screen "eProC - 09 - Estados PL_Diag" 1280x770, template "Template"
   Rectangle "Rectángulo_1" at 146,344 size 393x149
      Visibility <- "STOP_RUN"
   Button "Botón_2" at 352,429 size 144x40; TextOff 'Reset'
      on Click: SetBit("PL_Reset")
      Visibility <- "STOP_RUN"
   Button "Botón_1" at 192,429 size 144x40; TextOff 'Continuar'
      on Click: SetBit("PL_Continuar")
      Visibility <- "STOP_RUN"
   TextField "Campo de texto_17" at 165,356 size 351x73; Text 'Se ha detectado un reinicio del PLC. ¿Qué desea hacer con el ciclo de la Plegadora?'
      Visibility <- "STOP_RUN"
   Rectangle "Rectángulo_13" at 687,65 size 29x579
      Visibility <- "PL_S_1"
   Rectangle "Rectángulo_15" at 727,65 size 29x579
      Visibility <- "PL_S_2"
   Rectangle "Rectángulo_16" at 767,65 size 29x579
      Visibility <- "PL_S_9"
   Rectangle "Rectángulo_17" at 807,65 size 29x579
      Visibility <- "PL_S_3"
   Rectangle "Rectángulo_18" at 847,65 size 29x579
      Visibility <- "PL_S_4"
   Rectangle "Rectángulo_19" at 887,65 size 29x579
      Visibility <- "PL_S_10"
   Rectangle "Rectángulo_20" at 927,65 size 29x579
      Visibility <- "PL_S_5"
   Rectangle "Rectángulo_21" at 967,65 size 29x579
      Visibility <- "PL_S_11"
   Rectangle "Rectángulo_22" at 1007,65 size 29x579
      Visibility <- "PL_S_6"
   Rectangle "Rectángulo_23" at 647,65 size 29x579
      Visibility <- "PL_S_12"
   Circle "Círculo_2" at 78,143 size 450x450
      Appearance <- "PL_en_Ciclo"
   SymbolicIOField "Campo ES simbólico_1" at 109,310 size 387x69; TextOn '1'; TextOff '0'; TextList "Estados_PL"
      ProcessValue <- "PL_Estados"
   Polygon "Polígono_1" at 466,215 size 12x13
      Appearance <- "PL_en_Ciclo"
   Polygon "Polígono_2" at 520,333 size 8x12
      Appearance <- "PL_en_Ciclo"
   Polygon "Polígono_3" at 503,456 size 8x12
      Appearance <- "PL_en_Ciclo"
   Polygon "Polígono_4" at 401,559 size 14x10
      Appearance <- "PL_en_Ciclo"
   Polygon "Polígono_5" at 242,583 size 14x7
      Appearance <- "PL_en_Ciclo"
   Polygon "Polígono_6" at 124,503 size 10x13
      Appearance <- "PL_en_Ciclo"
   Polygon "Polígono_7" at 78,389 size 6x17
      Appearance <- "PL_en_Ciclo"
   Polygon "Polígono_8" at 94,269 size 7x14
      Appearance <- "PL_en_Ciclo"
   Polygon "Polígono_9" at 345,145 size 13x6
      Appearance <- "PL_en_Ciclo"
   Polygon "Polígono_10" at 186,169 size 12x9
      Appearance <- "PL_en_Ciclo"
   GraphicIOField "Campo ES gráfico_1" at 90,461 size 50x46; PictureList "Estado"
      ProcessValue <- "PL_S_11"
   GraphicIOField "Campo ES gráfico_2" at 55,345 size 50x46; PictureList "Estado"
      ProcessValue <- "PL_S_6"
   GraphicIOField "Campo ES gráfico_4" at 196,137 size 50x46; PictureList "Estado"
      ProcessValue <- "PL_S_1"
   GraphicIOField "Campo ES gráfico_5" at 196,555 size 50x46; PictureList "Estado"
      ProcessValue <- "PL_S_5"
   GraphicIOField "Campo ES gráfico_6" at 356,137 size 50x46; PictureList "Estado"
      ProcessValue <- "PL_S_2"
   GraphicIOField "Campo ES gráfico_7" at 356,554 size 50x46; PictureList "Estado"
      ProcessValue <- "PL_S_10"
   GraphicIOField "Campo ES gráfico_8" at 467,464 size 50x46; PictureList "Estado"
      ProcessValue <- "PL_S_4"
   GraphicIOField "Campo ES gráfico_9" at 466,226 size 50x46; PictureList "Estado"
      ProcessValue <- "PL_S_9"
   GraphicIOField "Campo ES gráfico_10" at 501,345 size 50x46; PictureList "Estado"
      ProcessValue <- "PL_S_3"
   SymbolicIOField "Campo ES simbólico_2" at 103,359 size 403x45; TextOn '1'; TextOff '0'; TextList "Transiciones_PL"
      ProcessValue <- "PL_Estados"
   Line "Línea_1" at 109,126 size 0x102
      Appearance <- "PL_en_Ciclo"
   Polygon "Polígono_11" at 106,213 size 7x15
      Appearance <- "PL_en_Ciclo"
   GraphicIOField "Campo ES gráfico_11" at 84,121 size 50x46; PictureList "Estado"
      ProcessValue <- "PL_S_0"
   GraphicIOField "Campo ES gráfico_3" at 86,226 size 50x46; PictureList "Estado"
      ProcessValue <- "PL_S_12"
   TextField "Campo de texto_1" at 31,36 size 300x29; Text 'Máquina de estados Plegadores'
   TextField "Campo de texto_15" at 372,147 size 16x25; Text '2'
   TextField "Campo de texto_16" at 482,236 size 16x25; Text '9'
   TextField "Campo de texto_13" at 518,355 size 16x25; Text '3'
   TextField "Campo de texto_24" at 483,474 size 16x25; Text '4'
   TextField "Campo de texto_26" at 366,564 size 30x25; Text '10'
   TextField "Campo de texto_27" at 211,565 size 19x25; Text '5'
   TextField "Campo de texto_28" at 100,471 size 30x25; Text '11'
   TextField "Campo de texto_29" at 70,355 size 15x25; Text '6'
   TextField "Campo de texto_30" at 96,236 size 31x25; Text '12'
   TextField "Campo de texto_31" at 212,147 size 16x25; Text '1'
   TextField "Campo de texto_32" at 100,131 size 16x25; Text '0'
   TextField "Campo de texto_2" at 1101,68 size 42x21; Text 'M10.3'
   TextField "Campo de texto_3" at 1147,92 size 50x21; Text 'M180.0'
   TextField "Campo de texto_4" at 1145,116 size 50x21; Text 'M180.1'
   TextField "Campo de texto_5" at 1170,140 size 50x21; Text 'M180.3'
   TextField "Campo de texto_6" at 1176,164 size 50x21; Text 'M180.4'
   TextField "Campo de texto_8" at 1138,212 size 96x21; Text 'DB11.DBX46.0'
   TextField "Campo de texto_14" at 1134,500 size 50x21; Text 'M170.5'
   TextField "Campo de texto_7" at 1134,524 size 50x21; Text 'M170.6'
   TextField "Campo de texto_9" at 1140,548 size 50x21; Text 'M170.7'
   TextField "Campo de texto_10" at 1147,572 size 50x21; Text 'M171.0'
   TextField "Campo de texto_11" at 1149,596 size 50x21; Text 'M171.1'
   TextField "Campo de texto_18" at 1130,620 size 50x21; Text 'M171.2'
   TextField "Campo de texto_22" at 1141,260 size 50x21; Text 'M165.0'
   TextField "Campo de texto_23" at 1148,284 size 50x21; Text 'M165.1'
   TextField "Campo de texto_12" at 1119,308 size 50x21; Text 'M165.2'
   TextField "Campo de texto_25" at 1125,332 size 50x21; Text 'M165.3'
   TextField "Campo de texto_19" at 1121,356 size 50x21; Text 'M165.4'
   TextField "Campo de texto_20" at 1125,380 size 50x21; Text 'M165.5'
   TextField "Campo de texto_21" at 1131,404 size 50x21; Text 'M165.6'
   TextField "Campo de texto_33" at 1136,428 size 50x21; Text 'M165.7'
   TextField "Campo de texto_34" at 1158,452 size 50x21; Text 'M166.0'
   TextField "Campo de texto_35" at 1164,476 size 50x21; Text 'M166.2'
   TextField "Campo de texto_36" at 1045,68 size 52x21; Text 'En Ciclo'
   TextField "Campo de texto_37" at 1045,92 size 98x21; Text 'Posición Espera'
   TextField "Campo de texto_38" at 1045,116 size 99x21; Text 'Posición Recep.'
   TextField "Campo de texto_39" at 1045,140 size 123x21; Text 'Posición Pleg. Patas'
   TextField "Campo de texto_40" at 1045,164 size 128x21; Text 'Posición Pleg. Techo'
   TextField "Campo de texto_41" at 1045,188 size 138x21; Text 'Posición Pleg. Entrega'
   TextField "Campo de texto_42" at 1045,212 size 91x21; Text 'Pieza Presente'
   TextField "Campo de texto_44" at 1045,500 size 86x21; Text 'Tenaza Arriba'
   TextField "Campo de texto_45" at 1045,524 size 86x21; Text 'Tenaza Abajo'
   TextField "Campo de texto_46" at 1045,548 size 93x21; Text 'Tenaza Abierta'
   TextField "Campo de texto_47" at 1045,572 size 99x21; Text 'Tenaza Cerrada'
   TextField "Campo de texto_48" at 1045,596 size 103x21; Text 'Tenaza Adelante'
   TextField "Campo de texto_49" at 1045,620 size 82x21; Text 'Tenaza Atrás'
   TextField "Campo de texto_53" at 1045,260 size 95x21; Text 'Alineadores ON'
   TextField "Campo de texto_54" at 1045,284 size 100x21; Text 'Alineadores OFF'
   TextField "Campo de texto_55" at 1045,308 size 71x21; Text 'Cepillos ON'
   TextField "Campo de texto_56" at 1045,332 size 76x21; Text 'Cepillos OFF'
   TextField "Campo de texto_57" at 1045,356 size 74x21; Text 'Prensas ON'
   TextField "Campo de texto_58" at 1045,380 size 79x21; Text 'Prensas OFF'
   TextField "Campo de texto_59" at 1045,404 size 85x21; Text 'Fijaciones ON'
   TextField "Campo de texto_60" at 1045,428 size 90x21; Text 'Fijaciones OFF'
   TextField "Campo de texto_61" at 1045,452 size 112x21; Text 'Plegado Patas ON'
   TextField "Campo de texto_62" at 1045,476 size 117x21; Text 'Plegado Techo ON'
   TextField "Campo de texto_43" at 1186,188 size 50x21; Text 'M180.5'
   GraphicIOField "Campo ES gráfico_13" at 969,210 size 24x24; PictureList "CheckBox"
      ProcessValue <- "Plegadora\Plegadora.PresenciaPieza"
   GraphicIOField "Campo ES gráfico_15" at 969,186 size 24x24; PictureList "CheckBox"
      ProcessValue <- "PL_En_Pos_Entrega"
   GraphicIOField "Campo ES gráfico_20" at 969,66 size 24x24; PictureList "CheckBox"
      ProcessValue <- "PL_en_Ciclo"
   GraphicIOField "Campo ES gráfico_27" at 929,522 size 24x24; PictureList "CheckBox"
      ProcessValue <- "PL_Tenaza_Abajo"
   GraphicIOField "Campo ES gráfico_29" at 929,474 size 24x24; PictureList "CheckBox"
      ProcessValue <- "PL_Plegador2_ON"
   GraphicIOField "Campo ES gráfico_32" at 929,402 size 24x24; PictureList "CheckBox"
      ProcessValue <- "PL_Fijaciones_SI"
   GraphicIOField "Campo ES gráfico_34" at 929,354 size 24x24; PictureList "CheckBox"
      ProcessValue <- "PL_Prensas_SI"
   GraphicIOField "Campo ES gráfico_39" at 929,210 size 24x24; PictureList "CheckBox"
      ProcessValue <- "Plegadora\Plegadora.PresenciaPieza"
   GraphicIOField "Campo ES gráfico_45" at 929,66 size 24x24; PictureList "CheckBox"
      ProcessValue <- "PL_en_Ciclo"
   GraphicIOField "Campo ES gráfico_46" at 929,570 size 24x24; PictureList "CheckBox"
      ProcessValue <- "PL_Tenaza_Cerrada"
   GraphicIOField "Campo ES gráfico_48" at 929,618 size 24x24; PictureList "CheckBox"
      ProcessValue <- "PL_Tenaza_Atrás"
   GraphicIOField "Campo ES gráfico_64" at 889,210 size 24x24; PictureList "CheckBox"
      ProcessValue <- "Plegadora\Plegadora.PresenciaPieza"
   GraphicIOField "Campo ES gráfico_66" at 889,162 size 24x24; PictureList "CheckBox"
      ProcessValue <- "PL_En_Pos_Pleg2"
   GraphicIOField "Campo ES gráfico_70" at 889,66 size 24x24; PictureList "CheckBox"
      ProcessValue <- "PL_en_Ciclo"
   GraphicIOField "Campo ES gráfico_77" at 849,522 size 24x24; PictureList "CheckBox"
      ProcessValue <- "PL_Tenaza_Abajo"
   GraphicIOField "Campo ES gráfico_80" at 849,450 size 24x24; PictureList "CheckBox"
      ProcessValue <- "PL_Plegador1_ON"
   GraphicIOField "Campo ES gráfico_82" at 849,402 size 24x24; PictureList "CheckBox"
      ProcessValue <- "PL_Fijaciones_SI"
   GraphicIOField "Campo ES gráfico_84" at 849,354 size 24x24; PictureList "CheckBox"
      ProcessValue <- "PL_Prensas_SI"
   GraphicIOField "Campo ES gráfico_89" at 849,210 size 24x24; PictureList "CheckBox"
      ProcessValue <- "Plegadora\Plegadora.PresenciaPieza"
   GraphicIOField "Campo ES gráfico_95" at 849,66 size 24x24; PictureList "CheckBox"
      ProcessValue <- "PL_en_Ciclo"
   GraphicIOField "Campo ES gráfico_96" at 849,570 size 24x24; PictureList "CheckBox"
      ProcessValue <- "PL_Tenaza_Cerrada"
   GraphicIOField "Campo ES gráfico_98" at 849,618 size 24x24; PictureList "CheckBox"
      ProcessValue <- "PL_Tenaza_Atrás"
   GraphicIOField "Campo ES gráfico_114" at 809,210 size 24x24; PictureList "CheckBox"
      ProcessValue <- "Plegadora\Plegadora.PresenciaPieza"
   GraphicIOField "Campo ES gráfico_117" at 809,138 size 24x24; PictureList "CheckBox"
      ProcessValue <- "PL_En_Pos_Pleg1"
   GraphicIOField "Campo ES gráfico_120" at 809,66 size 24x24; PictureList "CheckBox"
      ProcessValue <- "PL_en_Ciclo"
   GraphicIOField "Campo ES gráfico_127" at 769,522 size 24x24; PictureList "CheckBox"
      ProcessValue <- "PL_Tenaza_Abajo"
   GraphicIOField "Campo ES gráfico_131" at 769,426 size 24x24; PictureList "CheckBox"
      ProcessValue <- "PL_Fijaciones_No"
   GraphicIOField "Campo ES gráfico_133" at 769,378 size 24x24; PictureList "CheckBox"
      ProcessValue <- "PL_Prensas_No"
   GraphicIOField "Campo ES gráfico_135" at 769,330 size 24x24; PictureList "CheckBox"
      ProcessValue <- "PL_Cepillos_No"
   GraphicIOField "Campo ES gráfico_138" at 769,258 size 24x24; PictureList "CheckBox"
      ProcessValue <- "PL_Alineado_SI"
   GraphicIOField "Campo ES gráfico_139" at 769,210 size 24x24; PictureList "CheckBox"
      ProcessValue <- "Plegadora\Plegadora.PresenciaPieza"
   GraphicIOField "Campo ES gráfico_143" at 769,114 size 24x24; PictureList "CheckBox"
      ProcessValue <- "PL_En_Pos_Recepción"
   GraphicIOField "Campo ES gráfico_145" at 769,66 size 24x24; PictureList "CheckBox"
      ProcessValue <- "PL_en_Ciclo"
   GraphicIOField "Campo ES gráfico_148" at 769,618 size 24x24; PictureList "CheckBox"
      ProcessValue <- "PL_Tenaza_Atrás"
   GraphicIOField "Campo ES gráfico_151" at 729,546 size 24x24; PictureList "CheckBox"
      ProcessValue <- "PL_Tenaza_Abierta"
   GraphicIOField "Campo ES gráfico_152" at 729,522 size 24x24; PictureList "CheckBox"
      ProcessValue <- "PL_Tenaza_Abajo"
   GraphicIOField "Campo ES gráfico_170" at 729,66 size 24x24; PictureList "CheckBox"
      ProcessValue <- "PL_en_Ciclo"
   GraphicIOField "Campo ES gráfico_173" at 729,618 size 24x24; PictureList "CheckBox"
      ProcessValue <- "PL_Tenaza_Atrás"
   GraphicIOField "Campo ES gráfico_178" at 689,498 size 24x24; PictureList "CheckBox"
      ProcessValue <- "PL_Tenaza_Arriba"
   GraphicIOField "Campo ES gráfico_181" at 689,426 size 24x24; PictureList "CheckBox"
      ProcessValue <- "PL_Fijaciones_No"
   GraphicIOField "Campo ES gráfico_183" at 689,378 size 24x24; PictureList "CheckBox"
      ProcessValue <- "PL_Prensas_No"
   GraphicIOField "Campo ES gráfico_186" at 689,306 size 24x24; PictureList "CheckBox"
      ProcessValue <- "PL_Cepillos_SI"
   GraphicIOField "Campo ES gráfico_187" at 689,282 size 24x24; PictureList "CheckBox"
      ProcessValue <- "PL_Alineado_No"
   GraphicIOField "Campo ES gráfico_189" at 689,210 size 24x24; PictureList "CheckBox"
      ProcessValue <- "Plegadora\Plegadora.PresenciaPieza"
   GraphicIOField "Campo ES gráfico_193" at 689,114 size 24x24; PictureList "CheckBox"
      ProcessValue <- "PL_En_Pos_Recepción"
   GraphicIOField "Campo ES gráfico_195" at 689,66 size 24x24; PictureList "CheckBox"
      ProcessValue <- "PL_en_Ciclo"
   GraphicIOField "Campo ES gráfico_196" at 689,570 size 24x24; PictureList "CheckBox"
      ProcessValue <- "PL_Tenaza_Cerrada"
   GraphicIOField "Campo ES gráfico_197" at 689,594 size 24x24; PictureList "CheckBox"
      ProcessValue <- "PL_Tenaza_Adelante"
   GraphicIOField "Campo ES gráfico_214" at 649,210 size 24x24; PictureList "CheckBox"
      ProcessValue <- "Plegadora\Plegadora.PresenciaPieza"
   GraphicIOField "Campo ES gráfico_219" at 649,90 size 24x24; PictureList "CheckBox"
      ProcessValue <- "PL_En_Pos_Espera"
   GraphicIOField "Campo ES gráfico_220" at 649,66 size 24x24; PictureList "CheckBox"
      ProcessValue <- "PL_en_Ciclo"
   GraphicIOField "Campo ES gráfico_153" at 729,210 size 24x24; PictureList "CheckBox"
      ProcessValue <- "Plegadora\Plegadora.PresenciaPieza"
   GraphicIOField "Campo ES gráfico_53" at 1009,66 size 24x24; PictureList "CheckBox"
      ProcessValue <- "PL_en_Ciclo"
   TextField "Campo de texto_70" at 1160,236 size 96x21; Text 'DB11.DBX46.0'
   TextField "Campo de texto_71" at 1045,236 size 113x21; Text 'Sin Pieza Presente'
   GraphicIOField "Campo ES gráfico_12" at 1009,234 size 24x24; PictureList "CheckBox_Neg"
      ProcessValue <- "Plegadora\Plegadora.PresenciaPieza"
   Button "Botón_5" at 48,569 size 40x40; TextOff 'Vista Condiciones'; PictureOff "Gráfico_9"
      on Click: ActivateScreen("eProC - 09 - Estados PL", 0)
   Button "Botón_42" at 48,625 size 40x40; TextOff 'Vista Condiciones'; PictureOff "Gráfico_7"
      on Click: ActivateScreen("eProC - 09 - Estados PL_HW", 0)
   TextField "Campo de texto_50" at 249,678 size 130x18; Text 'DATOS PIEZA ACTUAL'
   TextField "Campo de texto_51" at 403,678 size 12x18; Text 'A'
   IOField "Champ E/S_24" at 414,675 size 53x25; FormatPattern 9999999
      ProcessValue <- "Plegadora\Plegadora.A"
      Appearance <- "Plegadora\Plegadora.PresenciaPieza"
   IOField "Champ E/S_25" at 483,675 size 53x25; FormatPattern 9999999
      ProcessValue <- "Plegadora\Plegadora.B"
      Appearance <- "Plegadora\Plegadora.PresenciaPieza"
   IOField "Champ E/S_26" at 554,675 size 53x24; FormatPattern 9999999
      ProcessValue <- "Plegadora\Plegadora.C"
      Appearance <- "Plegadora\Plegadora.PresenciaPieza"
   IOField "Champ E/S_27" at 629,675 size 53x25; FormatPattern 9999999
      ProcessValue <- "Plegadora\Plegadora.D"
      Appearance <- "Plegadora\Plegadora.PresenciaPieza"
   TextField "Campo de texto_52" at 472,678 size 11x18; Text 'B'
   TextField "Campo de texto_63" at 541,678 size 11x18; Text 'C'
   TextField "Campo de texto_64" at 616,678 size 12x18; Text 'D'
   Button "Botón_16" at 160,669 size 80x36; TextOff 'Borrar'; PictureOff "Borrar Pulsador"
      on Click: ResetBit("Plegadora\Plegadora.PresenciaPieza")
      Visibility <- "Plegadora\Plegadora.PresenciaPieza"
   Button "Botón_11" at 1224,27 size 40x37; TextOff 'Vista Condiciones'; PictureOff "Tool"; Authorization "Nivel 3"
      on Click: ActivateScreen("eProC - 11 Referencias F-PL", 0)
   Button "Template_Plantilla_Botón_5" at 789,715 size 150x53; TextOff 'PLEGADO'
      on Click: ActivateScreen("eProC - 09 - Estados PL", 0)
   TextField "Campo de texto_170" at 717,678 size 35x18; Text 'PL1-1'
   IOField "Champ E/S_162" at 752,675 size 51x25; FormatPattern s999999
      ProcessValue <- "Plegadora\Plegadora.PL1_1"
      Appearance <- "Plegadora\Plegadora.PresenciaPieza"
   IOField "Champ E/S_163" at 857,675 size 51x25; FormatPattern s999999
      ProcessValue <- "Plegadora\Plegadora.PL1_2"
      Appearance <- "Plegadora\Plegadora.PresenciaPieza"
   IOField "Champ E/S_164" at 962,675 size 51x24; FormatPattern s999999
      ProcessValue <- "Plegadora\Plegadora.PL2_1"
      Appearance <- "Plegadora\Plegadora.PresenciaPieza"
   IOField "Champ E/S_165" at 1060,675 size 51x25; FormatPattern s999999
      ProcessValue <- "Plegadora\Plegadora.PL2_2"
      Appearance <- "Plegadora\Plegadora.PresenciaPieza"
   TextField "Campo de texto_171" at 821,678 size 35x18; Text 'PL1-2'
   TextField "Campo de texto_172" at 925,678 size 35x18; Text 'PL2-1'
   TextField "Campo de texto_173" at 1023,678 size 35x18; Text 'PL2-2'

screen "eProC - 09 - Estados PL_HW" 1280x770, template "Template"
   GraphicIOField "Campo ES gráfico_7" at 255,205 size 757x290; PictureList "Pleg3"
      ProcessValue <- "Alarma_Plegador"
   Polygon "Polígono_2" at 289,278 size 725x83
      Visibility <- "Plegadora\Plegadora.PresenciaPieza"
   Circle "Cercle_9" at 614,250 size 8x8
      Appearance <- "30S2"
   Circle "Cercle_10" at 622,259 size 8x8
      Appearance <- "30S1"
   Circle "Cercle" at 604,253 size 8x8
      Appearance <- "30S4"
   Circle "Cercle_0" at 604,242 size 8x8
      Appearance <- "30S3"
   Circle "Cercle_11" at 442,264 size 8x8
      Appearance <- "32S1"
   Circle "Cercle_12" at 442,251 size 8x8
      Appearance <- "36S9"
   Circle "Cercle_13" at 442,236 size 8x8
      Appearance <- "32S2"
   Circle "Cercle_14" at 431,277 size 8x8
      Appearance <- "31S7b"
   Circle "Cercle_15" at 423,279 size 8x8
      Appearance <- "31S7"
   Circle "Cercle_18" at 436,285 size 8x8
      Appearance <- "30S7"
   Circle "Cercle_19" at 436,291 size 8x8
      Appearance <- "30S8"
   Circle "Cercle_20" at 415,308 size 8x8
      Appearance <- "23S5"
   Circle "Cercle_21" at 416,315 size 8x8
      Appearance <- "23S6"
   Circle "Cercle_22" at 454,361 size 8x8
      Appearance <- "31S8"
   Circle "Cercle_23" at 484,356 size 8x8
      Appearance <- "31S6"
   Circle "Cercle_24" at 484,321 size 8x8
      Appearance <- "31S5"
   Circle "Cercle_25" at 605,385 size 8x8
      Appearance <- "HommingPL1"
   Circle "Cercle_26" at 736,373 size 8x8
      Appearance <- "HommignPL2"
   Circle "Cercle_27" at 661,324 size 8x8
      Appearance <- "30S6"
   Circle "Cercle_28" at 676,300 size 8x8
      Appearance <- "30S5"
   Circle "Cercle_29" at 807,347 size 8x8
      Appearance <- "35S4"
   Circle "Cercle_30" at 831,323 size 8x8
      Appearance <- "35S2"
   Circle "Cercle_31" at 829,290 size 8x8
      Appearance <- "35S1"
   Circle "Cercle_32" at 883,270 size 8x8
      Appearance <- "35S3_0"
   Circle "Cercle_33" at 884,278 size 8x8
      Appearance <- "35S4"
   Circle "Cercle_34" at 821,266 size 8x8
      Appearance <- "36S8"
   Circle "Cercle_35" at 821,279 size 8x8
      Appearance <- "36S7"
   Circle "Cercle_36" at 812,254 size 8x8
      Appearance <- "35S8"
   Circle "Cercle_37" at 812,267 size 8x8
      Appearance <- "35S7"
   Circle "Cercle_38" at 862,240 size 8x8
      Appearance <- "36S2"
   Circle "Cercle_39" at 856,231 size 8x8
      Appearance <- "36S1"
   Circle "Cercle_40" at 830,246 size 8x8
      Appearance <- "36S5"
   Circle "Cercle_41" at 830,252 size 8x8
      Appearance <- "36S6"
   Circle "Cercle_42" at 815,222 size 8x8
      Appearance <- "35S3"
   Circle "Cercle_43" at 789,215 size 8x8
      Appearance <- "35S6"
   Circle "Cercle_45" at 790,246 size 8x8
      Appearance <- "35S5"
   Circle "Cercle_46" at 472,281 size 8x8
      Appearance <- "32S4"
   Circle "Cercle_47" at 470,295 size 8x8
      Appearance <- "32S3"
   Circle "Cercle_48" at 479,291 size 8x8
      Appearance <- "32S6"
   Circle "Cercle_49" at 477,305 size 8x8
      Appearance <- "32S5"
   TextField "Campo de texto_34" at 497,223 size 87x32; Text '30S3 - Tenaza Arriba'
   TextField "Campo de texto_35" at 501,178 size 87x32; Text '30S2 - Tenaza Atrás'
   TextField "Campo de texto_36" at 504,142 size 87x32; Text '30S1 - Tenaza Adelante'
   TextField "Campo de texto_37" at 497,260 size 87x32; Text '30S4 - Tenaza Abajo'
   TextField "Campo de texto_39" at 1004,467 size 99x18; Text '35S4 - PL2 Abajo'
   TextField "Campo de texto_40" at 735,507 size 126x18; Text '30S5 - Tenaza Abierta'
   TextField "Campo de texto_41" at 486,510 size 128x18; Text '30S6 - Tenaza Cerrada'
   TextField "Campo de texto_42" at 918,492 size 123x18; Text 'S16X20 - Homing PL2'
   TextField "Campo de texto_43" at 464,488 size 123x18; Text 'S16X20 - Homing PL1'
   TextField "Campo de texto_44" at 262,523 size 142x18; Text '31S6 - PL1 Fijación Abajo'
   TextField "Campo de texto_45" at 237,497 size 99x18; Text '31S8 - PL1 Abajo'
   TextField "Campo de texto_46" at 90,441 size 142x18; Text '31S5 - PL1 Fijación Arriba'
   TextField "Campo de texto_47" at 1036,443 size 118x18; Text '35S2 - Fijación Abajo'
   TextField "Campo de texto_48" at 1037,373 size 118x18; Text '35S1 - Fijación Arriba'
   TextField "Campo de texto_49" at 999,330 size 111x18; Text '36S4 - Alin. Y2 OFF'
   TextField "Campo de texto_50" at 999,305 size 107x18; Text '36S3 - Alin. Y2 ON'
   TextField "Campo de texto_51" at 975,226 size 108x18; Text '36S8 - Ext 2 Arriba'
   TextField "Campo de texto_52" at 975,243 size 108x18; Text '36S7 - Ext 2 Abajo'
   TextField "Campo de texto_53" at 655,262 size 108x18; Text '35S8 - Ext 1 Abajo'
   TextField "Campo de texto_54" at 655,246 size 108x18; Text '35S7 - Ext 1 Arriba'
   TextField "Campo de texto_55" at 1017,140 size 99x18; Text '36S1 - Alin. X ON'
   TextField "Campo de texto_56" at 1017,163 size 103x18; Text '36S2 - Alin. X OFF'
   TextField "Campo de texto_57" at 524,77 size 115x18; Text '35S6 - Prensa Arriba'
   TextField "Campo de texto_58" at 921,100 size 118x18; Text '36S5 - Cepillos Arriba'
   TextField "Campo de texto_59" at 935,117 size 118x18; Text '35S6 - Cepillos Abajo'
   TextField "Campo de texto_60" at 630,213 size 115x18; Text '35S5 - Prensa Abajo'
   TextField "Campo de texto_62" at 135,336 size 111x18; Text '23S6 - Alin. Y1 OFF'
   TextField "Campo de texto_63" at 140,318 size 107x18; Text '23S5 - Alin. Y1 ON'
   TextField "Campo de texto_64" at 169,170 size 115x18; Text '32S1 - Prensa Abajo'
   TextField "Campo de texto_65" at 141,145 size 143x18; Text '36S9 - Prensa Intermedia'
   TextField "Campo de texto_66" at 169,126 size 115x18; Text '32S2 - Prensa Arriba'
   TextField "Campo de texto_67" at 184,403 size 108x18; Text '32S5 - Ext 2 Abajo'
   TextField "Campo de texto_68" at 306,88 size 108x18; Text '32S6 - Ext 2 Arriba'
   TextField "Campo de texto_69" at 184,380 size 108x18; Text '32S3 - Ext 1 Abajo'
   TextField "Campo de texto_70" at 270,103 size 108x18; Text '32S4 - Ext 1 Arriba'
   TextField "Campo de texto_71" at 104,195 size 144x18; Text '31S7b - PL1 Arriba (Pata)'
   TextField "Campo de texto_72" at 148,215 size 99x18; Text '31S7 - PL1 Arriba'
   TextField "Campo de texto_75" at 127,271 size 118x18; Text '30S7 - Cepillos Arriba'
   TextField "Campo de texto_76" at 129,299 size 118x18; Text '30S8 - Cepillos Abajo'
   TextField "Campo de texto_77" at 887,59 size 99x18; Text '35S3 - PL2 Arriba'
   Circle "Cercle_50" at 807,223 size 8x8
      Appearance <- "35S3b"
   TextField "Campo de texto_78" at 907,76 size 144x18; Text '35S3b - PL2 Arriba (Pata)'
   Circle "Cercle_51" at 790,234 size 8x8
      Appearance <- "36S17"
   TextField "Campo de texto_79" at 491,99 size 150x18; Text '36S17 - Prensa Intermedia'
   Circle "Cercle_1" at 912,357 size 8x8
      Appearance <- "DI9_CU_PL"
   Circle "Cercle_2" at 365,401 size 8x8
      Appearance <- "DI8_CU_PL"
   TextField "Campo de texto_1" at 96,478 size 103x18; Text 'Fin de Carrera PL1'
   TextField "Campo de texto_2" at 1044,415 size 103x18; Text 'Fin de Carrera PL2'
   Circle "Cercle_3" at 375,268 size 8x8
      Appearance <- "21S5"
   Circle "Cercle_4" at 376,275 size 8x8
      Appearance <- "21S6"
   TextField "Campo de texto_3" at 129,252 size 110x18; Text '21S6 - Alin. X1 OFF'
   TextField "Campo de texto_4" at 134,234 size 106x18; Text '21S5 - Alin. X1 ON'
   Button "Botón_42" at 48,625 size 40x40; TextOff 'Vista Condiciones'; PictureOff "Gráfico_6"
      on Click: ActivateScreen("eProC - 09 - Estados PL", 0)
   Button "Botón_4" at 263,596 size 94x45; TextOff 'Plegador 1'
      on Press: SetTag("Selec_Pleg", 1)
      Visibility <- "MANU"
      Appearance <- "Selec_Pleg"
   Button "Botón_9" at 366,596 size 94x45; TextOff 'Plegador 2'
      on Press: SetTag("Selec_Pleg", 2)
      Visibility <- "MANU"
      Appearance <- "Selec_Pleg"
   Button "Botón_10" at 159,596 size 94x45; TextOff 'General'
      on Press: SetTag("Selec_Pleg", 3)
      Visibility <- "MANU"
      Appearance <- "Selec_Pleg"
   SymbolicIOField "Campo ES simbólico_3" at 734,569 size 230x29; TextOn '1'; TextOff '0'; TextList "SelecciónPlegadora"
      ProcessValue <- "Selec_Pleg"
      Visibility <- "Selec_Pleg"
   Button "Botón_6" at 730,596 size 69x33; TextOff 'Subir'
      on Press: SetTag("DB_OP.RC2", 18); SetBit("DB_OP.OP_SELMANU2")
      Visibility <- "Selec_Pleg"
      Appearance <- "DB_OP.RC2"
   Button "Botón_7" at 730,633 size 69x33; TextOff 'Bajar'
      on Press: SetTag("DB_OP.RC2", 19); SetBit("DB_OP.OP_SELMANU2")
      Visibility <- "Selec_Pleg"
      Appearance <- "DB_OP.RC2"
   Button "Botón_8" at 806,596 size 77x33; TextOff 'Avance'
      on Press: SetTag("DB_OP.RC2", 61); SetBit("DB_OP.OP_SELMANU2")
      Visibility <- "Selec_Pleg"
      Appearance <- "DB_OP.RC2"
   Button "Botón_11" at 806,633 size 77x33; TextOff 'Retroceso'
      on Press: SetTag("DB_OP.RC2", 62); SetBit("DB_OP.OP_SELMANU2")
      Visibility <- "Selec_Pleg"
      Appearance <- "DB_OP.RC2"
   Button "Botón_12" at 889,596 size 69x33; TextOff 'Bloquear'
      on Press: SetTag("DB_OP.RC2", 10); SetBit("DB_OP.OP_SELMANU2")
      Visibility <- "Selec_Pleg"
      Appearance <- "DB_OP.RC2"
   Button "Botón_13" at 889,633 size 69x33; TextOff 'Desbloquear'
      on Press: SetTag("DB_OP.RC2", 11); SetBit("DB_OP.OP_SELMANU2")
      Visibility <- "Selec_Pleg"
      Appearance <- "DB_OP.RC2"
   Button "Botón_14" at 979,633 size 85x33; TextOff 'Bajar Prensa'
      on Press: SetTag("DB_OP.RC2", 12); SetBit("DB_OP.OP_SELMANU2")
      Visibility <- "Selec_Pleg"
      Appearance <- "DB_OP.RC2"
   Button "Botón_15" at 979,596 size 85x33; TextOff 'Subir Prensa'
      on Press: SetTag("DB_OP.RC2", 13); SetBit("DB_OP.OP_SELMANU2")
      Visibility <- "Selec_Pleg"
      Appearance <- "DB_OP.RC2"
   Button "Botón_17" at 1071,633 size 85x33; TextOff 'Bajar Ext 1'
      on Press: SetTag("DB_OP.RC2", 14); SetBit("DB_OP.OP_SELMANU2")
      Visibility <- "Selec_Pleg"
      Appearance <- "DB_OP.RC2"
   Button "Botón_18" at 1071,596 size 85x33; TextOff 'Subir Ext 1'
      on Press: SetTag("DB_OP.RC2", 15); SetBit("DB_OP.OP_SELMANU2")
      Visibility <- "Selec_Pleg"
      Appearance <- "DB_OP.RC2"
   Button "Botón_19" at 1162,633 size 85x33; TextOff 'Bajar Ext 2'
      on Press: SetTag("DB_OP.RC2", 16); SetBit("DB_OP.OP_SELMANU2")
      Visibility <- "Selec_Pleg"
      Appearance <- "DB_OP.RC2"
   Button "Botón_20" at 1162,596 size 85x33; TextOff 'Subir Ext 2'
      on Press: SetTag("DB_OP.RC2", 17); SetBit("DB_OP.OP_SELMANU2")
      Visibility <- "Selec_Pleg"
      Appearance <- "DB_OP.RC2"
   Polyline "Línea poligonal_5" at 1025,674 size 69x11
      Visibility <- "Selec_Pleg"
   TextField "Campo de texto_19" at 1097,675 size 40x18; Text 'Prensa'
      Visibility <- "Selec_Pleg"
   Polyline "Línea poligonal_6" at 1140,674 size 69x11
      Visibility <- "Selec_Pleg"
   Button "Botón_21" at 730,596 size 69x33; TextOff 'Subir'
      on Press: SetTag("DB_OP.RC2", 28); SetBit("DB_OP.OP_SELMANU2")
      Visibility <- "Selec_Pleg"
      Appearance <- "DB_OP.RC2"
   Button "Botón_22" at 730,633 size 69x33; TextOff 'Bajar'
      on Press: SetTag("DB_OP.RC2", 29); SetBit("DB_OP.OP_SELMANU2")
      Visibility <- "Selec_Pleg"
      Appearance <- "DB_OP.RC2"
   Button "Botón_23" at 806,596 size 77x33; TextOff 'Avance'
      on Press: SetTag("DB_OP.RC2", 65); SetBit("DB_OP.OP_SELMANU2")
      Visibility <- "Selec_Pleg"
      Appearance <- "DB_OP.RC2"
   Button "Botón_24" at 806,633 size 77x33; TextOff 'Retroceso'
      on Press: SetTag("DB_OP.RC2", 66); SetBit("DB_OP.OP_SELMANU2")